   "Carrier_28_SpareSafetyInput(2_1)" AT %I1764.1 : Bool;   // SPARE SAFETY INPUT
   "Carrier_28_SpareSafetyInput(2_2)" AT %I1764.2 : Bool;   // SPARE SAFETY INPUT
   "Carrier_28_SpareSafetyInput(2_3)" AT %I1764.3 : Bool;   // SPARE SAFETY INPUT
   "Carrier_28_SpareSafetyInput(2_4)" AT %I1764.4 : Bool;   // SPARE SAFETY INPUT
   "Carrier_28_SpareSafetyInput(2_5)" AT %I1764.5 : Bool;   // SPARE SAFETY INPUT
   "Carrier_28_SpareSafetyInput(2_6)" AT %I1764.6 : Bool;   // SPARE SAFETY INPUT
   "Carrier_28_SpareSafetyInput(2_7)" AT %I1764.7 : Bool;   // SPARE SAFETY INPUT
   "Carrier_28_Slot3_SafetyOutput" AT %IW1675 : Word;   // SLOT 3 SAFETY OUTPUT WORD
   "Carrier_28_Crash_Detect_OK" AT %I1675.0 : Bool;   // CARRIER CRASH DETECT
   "Carrier_28_SpareSafetyOutput(3_1)" AT %I1675.1 : Bool;   // SPARE SAFETY OUTPUT
   "Carrier_28_SpareSafetyOutput(3_2)" AT %I1675.2 : Bool;   // SPARE SAFETY OUTPUT
   "Carrier_28_SpareSafetyOutput(3_3)" AT %I1675.3 : Bool;   // SPARE SAFETY OUTPUT
   "Carrier_28_SpareSafetyOutput(3_4)" AT %I1675.4 : Bool;   // SPARE SAFETY OUTPUT
   "Carrier_28_SpareSafetyOutput(3_5)" AT %I1675.5 : Bool;   // SPARE SAFETY OUTPUT
   "Carrier_28_SpareSafetyOutput(3_6)" AT %I1675.6 : Bool;   // SPARE SAFETY OUTPUT
   "Carrier_28_SpareSafetyOutput(3_7)" AT %I1675.7 : Bool;   // SPARE SAFETY OUTPUT
   "Carrier_28_Slot4_Input" AT %IW1766 : Word;   // SLOT 4 INPUT WORD
   "Carrier_28_480VPowerOn_MDCB1" AT %I1766.0 : Bool;   // 480 VAC POWER ON MDCB 1
   "Carrier_28_SpareInput(4_1)" AT %I1766.1 : Bool;   // SPARE INPUT
   "Carrier_28_SpareInput(4_2)" AT %I1766.2 : Bool;   // SPARE INPUT
   "Carrier_28_SitopSelectStatus" AT %I1766.3 : Bool;   // SITOP SELECT STATUS
   "Carrier_28_DCsupplyOnPSCB2" AT %I1766.4 : Bool;   // DC SUPPLY ON PSCB 2
   "Carrier_28_SpareInput(4_5)" AT %I1766.5 : Bool;   // SPARE INPUT
   "Carrier_28_SpareInput(4_6)" AT %I1766.6 : Bool;   // SPARE INPUT
   "Carrier_28_SpareInput(4_7)" AT %I1766.7 : Bool;   // SPARE INPUT
   "Carrier_28_PB1_ProdHoldLH" AT %I1767.0 : Bool;   // PB 1 PRODUCTION HOLD LH
   "Carrier_28_PB2_ResetLH" AT %I1767.1 : Bool;   // PB 2 RESET LH
   "Carrier_28_PB3_ProdHoldRH" AT %I1767.2 : Bool;   // PB 3 PRODUCTION HOLD RH
   "Carrier_28_PB4_ResetRH" AT %I1767.3 : Bool;   // PB 4 RESET RH
   "Carrier_28_SpareInput(4_14)" AT %I1767.4 : Bool;   // SPARE INPUT
   "Carrier_28_SpareInput(4_15)" AT %I1767.5 : Bool;   // SPARE INPUT
   "Carrier_28_SpareInput(4_16)" AT %I1767.6 : Bool;   // SPARE INPUT
   "Carrier_28_SpareInput(4_17)" AT %I1767.7 : Bool;   // SPARE INPUT
   "Carrier_28_Slot5_Output" AT %IW1768 : Word;   // SLOT 5 OUTPUT WORD
   "Carrier_28_IRD400_HMI_24VDC_ENABLE" AT %I1768.0 : Bool;   // IRD 400 PANEL HMI 24V DC POWER
   "Carrier_28_FaultLight_LH" AT %I1768.1 : Bool;   // FAULT LIGHT LH
   "Carrier_28_RunLight_LH" AT %I1768.2 : Bool;   // RUN LIGHT LH
   "Carrier_28_FaultLight_RH" AT %I1768.3 : Bool;   // FAULT LIGHT RH
   "Carrier_28_RunLight_RH" AT %I1768.4 : Bool;   // RUN LIGHT RH
   "Carrier_28_SpareOutput(5_5)" AT %I1768.5 : Bool;   // SPARE OUTPUT
   "Carrier_28_SpareOutput(5_6)" AT %I1768.6 : Bool;   // SPARE OUTPUT
   "Carrier_28_SpareOutput(5_7)" AT %I1768.7 : Bool;   // SPARE OUTPUT
   "Carrier_28_ActualSpeed" AT %IW1770 : Word;   // ACTUAL SPEED
   "Carrier_28_CarrierDriveAlarm" AT %IW1772 : Word;   // CARRIER DRIVE ALARM
   "Carrier_28_CarrierDriveWarning" AT %IW1774 : Word;   // CARRIER DRIVE WARNING
   "Carrier_29_Status" AT %IW1800 : Word;   // CARRIER STATUS WORD
   "Carrier_29_Status.0" AT %I1800.0 : Bool;   // HEARTBEAT
   "Carrier_29_Status.1" AT %I1800.1 : Bool;   // MANUAL
   "Carrier_29_Status.2" AT %I1800.2 : Bool;   // IN_AUTO
   "Carrier_29_Status.3" AT %I1800.3 : Bool;   // POSITIONING_COMPLETE
   "Carrier_29_Status.4" AT %I1800.4 : Bool;   // PRODUCTION HOLD
   "Carrier_29_Status.5" AT %I1800.5 : Bool;   // CARRIER MOVING FORWARD
   "Carrier_29_Status.6" AT %I1800.6 : Bool;   // CARRIER MOVING REVERSE
   "Carrier_29_Status.7" AT %I1800.7 : Bool;   // CARRIER FAULT
   "Carrier_29_Status.8" AT %I1801.0 : Bool;   // CRASH DETECT TRIPPED
   "Carrier_29_Status.9" AT %I1801.1 : Bool;
   "Carrier_29_Status.10" AT %I1801.2 : Bool;
   "Carrier_29_Status.11" AT %I1801.3 : Bool;
   "Carrier_29_Status.12" AT %I1801.4 : Bool;
   "Carrier_29_Status.13" AT %I1801.5 : Bool;
   "Carrier_29_Status.14" AT %I1801.6 : Bool;
   "Carrier_29_Status.15" AT %I1801.7 : Bool;
   "Carrier_29_SDCFaultCode" AT %IW1802 : Word;   // SDC FAULT CODE
   "Carrier_29_CarrierPosition" AT %ID1804 : DWord;   // CARRIER POSITION
   "Carrier_29_CarrierNumber" AT %IW1808 : Word;   // CARRIER NUMBER
   "Carrier_29_G120DControlWord" AT %IW1810 : Word;   // G120D_STW1_CONTROL
   "Carrier_29_G120DControlWord.0" AT %I1810.0 : Bool;   // Bit_00_ON
   "Carrier_29_G120DControlWord.1" AT %I1810.1 : Bool;   // Bit_01_AUS2_INH
   "Carrier_29_G120DControlWord.2" AT %I1810.2 : Bool;   // Bit_02_AUS3_STOP
   "Carrier_29_G120DControlWord.3" AT %I1810.3 : Bool;   // Bit_03_EN
   "Carrier_29_G120DControlWord.4" AT %I1810.4 : Bool;   // Bit_04_EN_RAMP
   "Carrier_29_G120DControlWord.5" AT %I1810.5 : Bool;   // Bit_05_START_RAMP
   "Carrier_29_G120DControlWord.6" AT %I1810.6 : Bool;   // Bit_06_SETPOINT
   "Carrier_29_G120DControlWord.7" AT %I1810.7 : Bool;   // Bit_07_RESET
   "Carrier_29_G120DControlWord.8" AT %I1811.0 : Bool;   // Bit_08_JOG_R
   "Carrier_29_G120DControlWord.9" AT %I1811.1 : Bool;   // Bit_09_JOG_L
   "Carrier_29_G120DControlWord.10" AT %I1811.2 : Bool;   // Bit_10_CONTR_PLC
   "Carrier_29_G120DControlWord.11" AT %I1811.3 : Bool;   // Bit_11_REVERSE
   "Carrier_29_G120DControlWord.12" AT %I1811.4 : Bool;   // Bit_12_BRAKE_RELEASE
   "Carrier_29_G120DControlWord.13" AT %I1811.5 : Bool;   // Bit_13_DDS
   "Carrier_29_G120DControlWord.14" AT %I1811.6 : Bool;   // Bit_14_DO0
   "Carrier_29_G120DControlWord.15" AT %I1811.7 : Bool;   // Bit_15_DO1
   "Carrier_29_G120DStatusWord" AT %IW1812 : Word;   // G120D_ZSW1_STATUS
   "Carrier_29_G120DStatusWord.0" AT %I1812.0 : Bool;   // Bit_00_READY_RUN
   "Carrier_29_G120DStatusWord.1" AT %I1812.1 : Bool;   // Bit_01_READY_ON
   "Carrier_29_G120DStatusWord.2" AT %I1812.2 : Bool;   // Bit_02_ENABLE
   "Carrier_29_G120DStatusWord.3" AT %I1812.3 : Bool;   // Bit_03_FAULT
   "Carrier_29_G120DStatusWord.4" AT %I1812.4 : Bool;   // Bit_04_OFF2
   "Carrier_29_G120DStatusWord.5" AT %I1812.5 : Bool;   // Bit_05_OFF3
   "Carrier_29_G120DStatusWord.6" AT %I1812.6 : Bool;   // Bit_06_LOCK_OUT
   "Carrier_29_G120DStatusWord.7" AT %I1812.7 : Bool;   // Bit_07_WARN
   "Carrier_29_G120DStatusWord.8" AT %I1813.0 : Bool;   // Bit_08_NO_DEVIATION
   "Carrier_29_G120DStatusWord.9" AT %I1813.1 : Bool;   // Bit_09_CONTR_PLC
   "Carrier_29_G120DStatusWord.10" AT %I1813.2 : Bool;   // Bit_10_F_MAX
   "Carrier_29_G120DStatusWord.11" AT %I1813.3 : Bool;   // Bit_11_LIMIT_REACHED
   "Carrier_29_G120DStatusWord.12" AT %I1813.4 : Bool;   // Bit_12_BRAKE_OPEN
   "Carrier_29_G120DStatusWord.13" AT %I1813.5 : Bool;   // Bit_13_NO_OVERTEMP
   "Carrier_29_G120DStatusWord.14" AT %I1813.6 : Bool;   // Bit_14_CW_CCW
   "Carrier_29_G120DStatusWord.15" AT %I1813.7 : Bool;   // Bit_15_OVERL
   "Carrier_29_Slot2_Input" AT %IW1814 : Word;   // SLOT 2 INPUT WORD
   "Carrier_29_CrashDetectSW" AT %I1814.0 : Bool;   // CRASH DETECT SW
   "Carrier_29_SpareSafetyInput(2_1)" AT %I1814.1 : Bool;   // SPARE SAFETY INPUT
   "Carrier_29_SpareSafetyInput(2_2)" AT %I1814.2 : Bool;   // SPARE SAFETY INPUT
   "Carrier_29_SpareSafetyInput(2_3)" AT %I1814.3 : Bool;   // SPARE SAFETY INPUT
   "Carrier_29_SpareSafetyInput(2_4)" AT %I1814.4 : Bool;   // SPARE SAFETY INPUT
   "Carrier_29_SpareSafetyInput(2_5)" AT %I1814.5 : Bool;   // SPARE SAFETY INPUT
   "Carrier_29_SpareSafetyInput(2_6)" AT %I1814.6 : Bool;   // SPARE SAFETY INPUT
   "Carrier_29_SpareSafetyInput(2_7)" AT %I1814.7 : Bool;   // SPARE SAFETY INPUT
   "Carrier_29_Slot3_SafetyOutput" AT %IW1815 : Word;   // SLOT 3 SAFETY OUTPUT WORD
   "Carrier_29_Crash_Detect_OK" AT %I1815.0 : Bool;   // CARRIER CRASH DETECT
   "Carrier_29_SpareSafetyOutput(3_1)" AT %I1815.1 : Bool;   // SPARE SAFETY OUTPUT
   "Carrier_29_SpareSafetyOutput(3_2)" AT %I1815.2 : Bool;   // SPARE SAFETY OUTPUT
   "Carrier_29_SpareSafetyOutput(3_3)" AT %I1815.3 : Bool;   // SPARE SAFETY OUTPUT
   "Carrier_29_SpareSafetyOutput(3_4)" AT %I1815.4 : Bool;   // SPARE SAFETY OUTPUT
   "Carrier_29_SpareSafetyOutput(3_5)" AT %I1815.5 : Bool;   // SPARE SAFETY OUTPUT
   "Carrier_29_SpareSafetyOutput(3_6)" AT %I1815.6 : Bool;   // SPARE SAFETY OUTPUT
   "Carrier_29_SpareSafetyOutput(3_7)" AT %I1815.7 : Bool;   // SPARE SAFETY OUTPUT
   "Carrier_29_Slot4_Input" AT %IW1816 : Word;   // SLOT 4 INPUT WORD
   "Carrier_29_480VPowerOn_MDCB1" AT %I1816.0 : Bool;   // 480 VAC POWER ON MDCB 1
   "Carrier_29_SpareInput(4_1)" AT %I1816.1 : Bool;   // SPARE INPUT
   "Carrier_29_SpareInput(4_2)" AT %I1816.2 : Bool;   // SPARE INPUT
   "Carrier_29_SitopSelectStatus" AT %I1816.3 : Bool;   // SITOP SELECT STATUS
   "Carrier_29_DCsupplyOnPSCB2" AT %I1816.4 : Bool;   // DC SUPPLY ON PSCB 2
   "Carrier_29_SpareInput(4_5)" AT %I1816.5 : Bool;   // SPARE INPUT
   "Carrier_29_SpareInput(4_6)" AT %I1816.6 : Bool;   // SPARE INPUT
   "Carrier_29_SpareInput(4_7)" AT %I1816.7 : Bool;   // SPARE INPUT
   "Carrier_29_PB1_ProdHoldLH" AT %I1817.0 : Bool;   // PB 1 PRODUCTION HOLD LH
   "Carrier_29_PB2_ResetLH" AT %I1817.1 : Bool;   // PB 2 RESET LH
   "Carrier_29_PB3_ProdHoldRH" AT %I1817.2 : Bool;   // PB 3 PRODUCTION HOLD RH
   "Carrier_29_PB4_ResetRH" AT %I1817.3 : Bool;   // PB 4 RESET RH
   "Carrier_29_SpareInput(4_14)" AT %I1817.4 : Bool;   // SPARE INPUT
   "Carrier_29_SpareInput(4_15)" AT %I1817.5 : Bool;   // SPARE INPUT
   "Carrier_29_SpareInput(4_16)" AT %I1817.6 : Bool;   // SPARE INPUT
   "Carrier_29_SpareInput(4_17)" AT %I1817.7 : Bool;   // SPARE INPUT
   "Carrier_29_Slot5_Output" AT %IW1818 : Word;   // SLOT 5 OUTPUT WORD
   "Carrier_29_IRD400_HMI_24VDC_ENABLE" AT %I1818.0 : Bool;   // IRD 400 PANEL HMI 24V DC POWER
   "Carrier_29_FaultLight_LH" AT %I1818.1 : Bool;   // FAULT LIGHT LH
   "Carrier_29_RunLight_LH" AT %I1818.2 : Bool;   // RUN LIGHT LH
   "Carrier_29_FaultLight_RH" AT %I1818.3 : Bool;   // FAULT LIGHT RH
   "Carrier_29_RunLight_RH" AT %I1818.4 : Bool;   // RUN LIGHT RH
   "Carrier_29_SpareOutput(5_5)" AT %I1818.5 : Bool;   // SPARE OUTPUT
   "Carrier_29_SpareOutput(5_6)" AT %I1818.6 : Bool;   // SPARE OUTPUT
   "Carrier_29_SpareOutput(5_7)" AT %I1818.7 : Bool;   // SPARE OUTPUT
   "Carrier_29_ActualSpeed" AT %IW1820 : Word;   // ACTUAL SPEED
   "Carrier_29_CarrierDriveAlarm" AT %IW1822 : Word;   // CARRIER DRIVE ALARM
   "Carrier_29_CarrierDriveWarning" AT %IW1824 : Word;   // CARRIER DRIVE WARNING
   "Carrier_30_Status" AT %IW1850 : Word;   // CARRIER STATUS WORD
   "Carrier_30_Status.0" AT %I1850.0 : Bool;   // HEARTBEAT
   "Carrier_30_Status.1" AT %I1850.1 : Bool;   // MANUAL
   "Carrier_30_Status.2" AT %I1850.2 : Bool;   // IN_AUTO
   "Carrier_30_Status.3" AT %I1850.3 : Bool;   // POSITIONING_COMPLETE
   "Carrier_30_Status.4" AT %I1850.4 : Bool;   // PRODUCTION HOLD
   "Carrier_30_Status.5" AT %I1850.5 : Bool;   // CARRIER MOVING FORWARD
   "Carrier_30_Status.6" AT %I1850.6 : Bool;   // CARRIER MOVING REVERSE
   "Carrier_30_Status.7" AT %I1850.7 : Bool;   // CARRIER FAULT
   "Carrier_30_Status.8" AT %I1851.0 : Bool;   // CRASH DETECT TRIPPED
   "Carrier_30_Status.9" AT %I1851.1 : Bool;
   "Carrier_30_Status.10" AT %I1851.2 : Bool;
   "Carrier_30_Status.11" AT %I1851.3 : Bool;
   "Carrier_30_Status.12" AT %I1851.4 : Bool;
   "Carrier_30_Status.13" AT %I1851.5 : Bool;
   "Carrier_30_Status.14" AT %I1851.6 : Bool;
   "Carrier_30_Status.15" AT %I1851.7 : Bool;
   "Carrier_30_SDCFaultCode" AT %IW1852 : Word;   // SDC FAULT CODE
   "Carrier_30_CarrierPosition" AT %ID1854 : DWord;   // CARRIER POSITION
   "Carrier_30_CarrierNumber" AT %IW1858 : Word;   // CARRIER NUMBER
   "Carrier_30_G120DControlWord" AT %IW1860 : Word;   // G120D_STW1_CONTROL
   "Carrier_30_G120DControlWord.0" AT %I1860.0 : Bool;   // Bit_00_ON
   "Carrier_30_G120DControlWord.1" AT %I1860.1 : Bool;   // Bit_01_AUS2_INH
   "Carrier_30_G120DControlWord.2" AT %I1860.2 : Bool;   // Bit_02_AUS3_STOP
   "Carrier_30_G120DControlWord.3" AT %I1860.3 : Bool;   // Bit_03_EN
   "Carrier_30_G120DControlWord.4" AT %I1860.4 : Bool;   // Bit_04_EN_RAMP
   "Carrier_30_G120DControlWord.5" AT %I1860.5 : Bool;   // Bit_05_START_RAMP
   "Carrier_30_G120DControlWord.6" AT %I1860.6 : Bool;   // Bit_06_SETPOINT
   "Carrier_30_G120DControlWord.7" AT %I1860.7 : Bool;   // Bit_07_RESET
   "Carrier_30_G120DControlWord.8" AT %I1861.0 : Bool;   // Bit_08_JOG_R
   "Carrier_30_G120DControlWord.9" AT %I1861.1 : Bool;   // Bit_09_JOG_L
   "Carrier_30_G120DControlWord.10" AT %I1861.2 : Bool;   // Bit_10_CONTR_PLC
   "Carrier_30_G120DControlWord.11" AT %I1861.3 : Bool;   // Bit_11_REVERSE
   "Carrier_30_G120DControlWord.12" AT %I1861.4 : Bool;   // Bit_12_BRAKE_RELEASE
   "Carrier_30_G120DControlWord.13" AT %I1861.5 : Bool;   // Bit_13_DDS
   "Carrier_30_G120DControlWord.14" AT %I1861.6 : Bool;   // Bit_14_DO0
   "Carrier_30_G120DControlWord.15" AT %I1861.7 : Bool;   // Bit_15_DO1
   "Carrier_30_G120DStatusWord" AT %IW1862 : Word;   // G120D_ZSW1_STATUS
   "Carrier_30_G120DStatusWord.0" AT %I1862.0 : Bool;   // Bit_00_READY_RUN
   "Carrier_30_G120DStatusWord.1" AT %I1862.1 : Bool;   // Bit_01_READY_ON
   "Carrier_30_G120DStatusWord.2" AT %I1862.2 : Bool;   // Bit_02_ENABLE
   "Carrier_30_G120DStatusWord.3" AT %I1862.3 : Bool;   // Bit_03_FAULT
   "Carrier_30_G120DStatusWord.4" AT %I1862.4 : Bool;   // Bit_04_OFF2
   "Carrier_30_G120DStatusWord.5" AT %I1862.5 : Bool;   // Bit_05_OFF3
   "Carrier_30_G120DStatusWord.6" AT %I1862.6 : Bool;   // Bit_06_LOCK_OUT
   "Carrier_30_G120DStatusWord.7" AT %I1862.7 : Bool;   // Bit_07_WARN
   "Carrier_30_G120DStatusWord.8" AT %I1863.0 : Bool;   // Bit_08_NO_DEVIATION
   "Carrier_30_G120DStatusWord.9" AT %I1863.1 : Bool;   // Bit_09_CONTR_PLC
   "Carrier_30_G120DStatusWord.10" AT %I1863.2 : Bool;   // Bit_10_F_MAX
   "Carrier_30_G120DStatusWord.11" AT %I1863.3 : Bool;   // Bit_11_LIMIT_REACHED
   "Carrier_30_G120DStatusWord.12" AT %I1863.4 : Bool;   // Bit_12_BRAKE_OPEN
   "Carrier_30_G120DStatusWord.13" AT %I1863.5 : Bool;   // Bit_13_NO_OVERTEMP
   "Carrier_30_G120DStatusWord.14" AT %I1863.6 : Bool;   // Bit_14_CW_CCW
   "Carrier_30_G120DStatusWord.15" AT %I1863.7 : Bool;   // Bit_15_OVERL
   "Carrier_30_Slot2_Input" AT %IW1864 : Word;   // SLOT 2 INPUT WORD
   "Carrier_30_CrashDetectSW" AT %I1864.0 : Bool;   // CRASH DETECT SW
   "Carrier_30_SpareSafetyInput(2_1)" AT %I1864.1 : Bool;   // SPARE SAFETY INPUT
   "Carrier_30_SpareSafetyInput(2_2)" AT %I1864.2 : Bool;   // SPARE SAFETY INPUT
   "Carrier_30_SpareSafetyInput(2_3)" AT %I1864.3 : Bool;   // SPARE SAFETY INPUT
   "Carrier_30_SpareSafetyInput(2_4)" AT %I1864.4 : Bool;   // SPARE SAFETY INPUT
   "Carrier_30_SpareSafetyInput(2_5)" AT %I1864.5 : Bool;   // SPARE SAFETY INPUT
   "Carrier_30_SpareSafetyInput(2_6)" AT %I1864.6 : Bool;   // SPARE SAFETY INPUT
   "Carrier_30_SpareSafetyInput(2_7)" AT %I1864.7 : Bool;   // SPARE SAFETY INPUT
   "Carrier_30_Slot3_SafetyOutput" AT %IW1685 : Word;   // SLOT 3 SAFETY OUTPUT WORD
   "Carrier_30_Crash_Detect_OK" AT %I1685.0 : Bool;   // CARRIER CRASH DETECT
   "Carrier_30_SpareSafetyOutput(3_1)" AT %I1685.1 : Bool;   // SPARE SAFETY OUTPUT
   "Carrier_30_SpareSafetyOutput(3_2)" AT %I1685.2 : Bool;   // SPARE SAFETY OUTPUT
   "Carrier_30_SpareSafetyOutput(3_3)" AT %I1685.3 : Bool;   // SPARE SAFETY OUTPUT
   "Carrier_30_SpareSafetyOutput(3_4)" AT %I1685.4 : Bool;   // SPARE SAFETY OUTPUT
   "Carrier_30_SpareSafetyOutput(3_5)" AT %I1685.5 : Bool;   // SPARE SAFETY OUTPUT
   "Carrier_30_SpareSafetyOutput(3_6)" AT %I1685.6 : Bool;   // SPARE SAFETY OUTPUT
   "Carrier_30_SpareSafetyOutput(3_7)" AT %I1685.7 : Bool;   // SPARE SAFETY OUTPUT
   "Carrier_30_Slot4_Input" AT %IW1866 : Word;   // SLOT 4 INPUT WORD
   "Carrier_30_480VPowerOn_MDCB1" AT %I1866.0 : Bool;   // 480 VAC POWER ON MDCB 1
   "Carrier_30_SpareInput(4_1)" AT %I1866.1 : Bool;   // SPARE INPUT
   "Carrier_30_SpareInput(4_2)" AT %I1866.2 : Bool;   // SPARE INPUT
   "Carrier_30_SitopSelectStatus" AT %I1866.3 : Bool;   // SITOP SELECT STATUS
   "Carrier_30_DCsupplyOnPSCB2" AT %I1866.4 : Bool;   // DC SUPPLY ON PSCB 2
   "Carrier_30_SpareInput(4_5)" AT %I1866.5 : Bool;   // SPARE INPUT
   "Carrier_30_SpareInput(4_6)" AT %I1866.6 : Bool;   // SPARE INPUT
   "Carrier_30_SpareInput(4_7)" AT %I1866.7 : Bool;   // SPARE INPUT
   "Carrier_30_PB1_ProdHoldLH" AT %I1867.0 : Bool;   // PB 1 PRODUCTION HOLD LH
   "Carrier_30_PB2_ResetLH" AT %I1867.1 : Bool;   // PB 2 RESET LH
   "Carrier_30_PB3_ProdHoldRH" AT %I1867.2 : Bool;   // PB 3 PRODUCTION HOLD RH
   "Carrier_30_PB4_ResetRH" AT %I1867.3 : Bool;   // PB 4 RESET RH
   "Carrier_30_SpareInput(4_14)" AT %I1867.4 : Bool;   // SPARE INPUT
   "Carrier_30_SpareInput(4_15)" AT %I1867.5 : Bool;   // SPARE INPUT
   "Carrier_30_SpareInput(4_16)" AT %I1867.6 : Bool;   // SPARE INPUT
   "Carrier_30_SpareInput(4_17)" AT %I1867.7 : Bool;   // SPARE INPUT
   "Carrier_30_Slot5_Output" AT %IW1868 : Word;   // SLOT 5 OUTPUT WORD
   "Carrier_30_IRD400_HMI_24VDC_ENABLE" AT %I1868.0 : Bool;   // IRD 400 PANEL HMI 24V DC POWER
   "Carrier_30_FaultLight_LH" AT %I1868.1 : Bool;   // FAULT LIGHT LH
   "Carrier_30_RunLight_LH" AT %I1868.2 : Bool;   // RUN LIGHT LH
   "Carrier_30_FaultLight_RH" AT %I1868.3 : Bool;   // FAULT LIGHT RH
   "Carrier_30_RunLight_RH" AT %I1868.4 : Bool;   // RUN LIGHT RH
   "Carrier_30_SpareOutput(5_5)" AT %I1868.5 : Bool;   // SPARE OUTPUT
   "Carrier_30_SpareOutput(5_6)" AT %I1868.6 : Bool;   // SPARE OUTPUT
   "Carrier_30_SpareOutput(5_7)" AT %I1868.7 : Bool;   // SPARE OUTPUT
   "Carrier_30_ActualSpeed" AT %IW1870 : Word;   // ACTUAL SPEED
   "Carrier_30_CarrierDriveAlarm" AT %IW1872 : Word;   // CARRIER DRIVE ALARM
   "Carrier_30_CarrierDriveWarning" AT %IW1874 : Word;   // CARRIER DRIVE WARNING
   "Carrier_31_Status" AT %IW1900 : Word;   // CARRIER STATUS WORD
   "Carrier_31_Status.0" AT %I1900.0 : Bool;   // HEARTBEAT
   "Carrier_31_Status.1" AT %I1900.1 : Bool;   // MANUAL
   "Carrier_31_Status.2" AT %I1900.2 : Bool;   // IN_AUTO
   "Carrier_31_Status.3" AT %I1900.3 : Bool;   // POSITIONING_COMPLETE
   "Carrier_31_Status.4" AT %I1900.4 : Bool;   // PRODUCTION HOLD
   "Carrier_31_Status.5" AT %I1900.5 : Bool;   // CARRIER MOVING FORWARD
   "Carrier_31_Status.6" AT %I1900.6 : Bool;   // CARRIER MOVING REVERSE
   "Carrier_31_Status.7" AT %I1900.7 : Bool;   // CARRIER FAULT
   "Carrier_31_Status.8" AT %I1901.0 : Bool;   // CRASH DETECT TRIPPED
   "Carrier_31_Status.9" AT %I1901.1 : Bool;
   "Carrier_31_Status.10" AT %I1901.2 : Bool;
   "Carrier_31_Status.11" AT %I1901.3 : Bool;
   "Carrier_31_Status.12" AT %I1901.4 : Bool;
   "Carrier_31_Status.13" AT %I1901.5 : Bool;
   "Carrier_31_Status.14" AT %I1901.6 : Bool;
   "Carrier_31_Status.15" AT %I1901.7 : Bool;
   "Carrier_31_SDCFaultCode" AT %IW1902 : Word;   // SDC FAULT CODE
   "Carrier_31_CarrierPosition" AT %ID1904 : DWord;   // CARRIER POSITION
   "Carrier_31_CarrierNumber" AT %IW1908 : Word;   // CARRIER NUMBER
   "Carrier_31_G120DControlWord" AT %IW1910 : Word;   // G120D_STW1_CONTROL
   "Carrier_31_G120DControlWord.0" AT %I1910.0 : Bool;   // Bit_00_ON
   "Carrier_31_G120DControlWord.1" AT %I1910.1 : Bool;   // Bit_01_AUS2_INH
   "Carrier_31_G120DControlWord.2" AT %I1910.2 : Bool;   // Bit_02_AUS3_STOP
   "Carrier_31_G120DControlWord.3" AT %I1910.3 : Bool;   // Bit_03_EN
   "Carrier_31_G120DControlWord.4" AT %I1910.4 : Bool;   // Bit_04_EN_RAMP
   "Carrier_31_G120DControlWord.5" AT %I1910.5 : Bool;   // Bit_05_START_RAMP
   "Carrier_31_G120DControlWord.6" AT %I1910.6 : Bool;   // Bit_06_SETPOINT
   "Carrier_31_G120DControlWord.7" AT %I1910.7 : Bool;   // Bit_07_RESET
   "Carrier_31_G120DControlWord.8" AT %I1911.0 : Bool;   // Bit_08_JOG_R
   "Carrier_31_G120DControlWord.9" AT %I1911.1 : Bool;   // Bit_09_JOG_L
   "Carrier_31_G120DControlWord.10" AT %I1911.2 : Bool;   // Bit_10_CONTR_PLC
   "Carrier_31_G120DControlWord.11" AT %I1911.3 : Bool;   // Bit_11_REVERSE
   "Carrier_31_G120DControlWord.12" AT %I1911.4 : Bool;   // Bit_12_BRAKE_RELEASE
   "Carrier_31_G120DControlWord.13" AT %I1911.5 : Bool;   // Bit_13_DDS
   "Carrier_31_G120DControlWord.14" AT %I1911.6 : Bool;   // Bit_14_DO0
   "Carrier_31_G120DControlWord.15" AT %I1911.7 : Bool;   // Bit_15_DO1
   "Carrier_31_G120DStatusWord" AT %IW1912 : Word;   // G120D_ZSW1_STATUS
   "Carrier_31_G120DStatusWord.0" AT %I1912.0 : Bool;   // Bit_00_READY_RUN
   "Carrier_31_G120DStatusWord.1" AT %I1912.1 : Bool;   // Bit_01_READY_ON
   "Carrier_31_G120DStatusWord.2" AT %I1912.2 : Bool;   // Bit_02_ENABLE
   "Carrier_31_G120DStatusWord.3" AT %I1912.3 : Bool;   // Bit_03_FAULT
   "Carrier_31_G120DStatusWord.4" AT %I1912.4 : Bool;   // Bit_04_OFF2
   "Carrier_31_G120DStatusWord.5" AT %I1912.5 : Bool;   // Bit_05_OFF3
   "Carrier_31_G120DStatusWord.6" AT %I1912.6 : Bool;   // Bit_06_LOCK_OUT
   "Carrier_31_G120DStatusWord.7" AT %I1912.7 : Bool;   // Bit_07_WARN
   "Carrier_31_G120DStatusWord.8" AT %I1913.0 : Bool;   // Bit_08_NO_DEVIATION
   "Carrier_31_G120DStatusWord.9" AT %I1913.1 : Bool;   // Bit_09_CONTR_PLC
   "Carrier_31_G120DStatusWord.10" AT %I1913.2 : Bool;   // Bit_10_F_MAX
   "Carrier_31_G120DStatusWord.11" AT %I1913.3 : Bool;   // Bit_11_LIMIT_REACHED
   "Carrier_31_G120DStatusWord.12" AT %I1913.4 : Bool;   // Bit_12_BRAKE_OPEN
   "Carrier_31_G120DStatusWord.13" AT %I1913.5 : Bool;   // Bit_13_NO_OVERTEMP
   "Carrier_31_G120DStatusWord.14" AT %I1913.6 : Bool;   // Bit_14_CW_CCW
   "Carrier_31_G120DStatusWord.15" AT %I1913.7 : Bool;   // Bit_15_OVERL
   "Carrier_31_Slot2_Input" AT %IW1914 : Word;   // SLOT 2 INPUT WORD
   "Carrier_31_CrashDetectSW" AT %I1914.0 : Bool;   // CRASH DETECT SW
   "Carrier_31_SpareSafetyInput(2_1)" AT %I1914.1 : Bool;   // SPARE SAFETY INPUT
   "Carrier_31_SpareSafetyInput(2_2)" AT %I1914.2 : Bool;   // SPARE SAFETY INPUT
   "Carrier_31_SpareSafetyInput(2_3)" AT %I1914.3 : Bool;   // SPARE SAFETY INPUT
   "Carrier_31_SpareSafetyInput(2_4)" AT %I1914.4 : Bool;   // SPARE SAFETY INPUT
   "Carrier_31_SpareSafetyInput(2_5)" AT %I1914.5 : Bool;   // SPARE SAFETY INPUT
   "Carrier_31_SpareSafetyInput(2_6)" AT %I1914.6 : Bool;   // SPARE SAFETY INPUT
   "Carrier_31_SpareSafetyInput(2_7)" AT %I1914.7 : Bool;   // SPARE SAFETY INPUT
   "Carrier_31_Slot3_SafetyOutput" AT %IW1915 : Word;   // SLOT 3 SAFETY OUTPUT WORD
   "Carrier_31_Crash_Detect_OK" AT %I1915.0 : Bool;   // CARRIER CRASH DETECT
   "Carrier_31_SpareSafetyOutput(3_1)" AT %I1915.1 : Bool;   // SPARE SAFETY OUTPUT
   "Carrier_31_SpareSafetyOutput(3_2)" AT %I1915.2 : Bool;   // SPARE SAFETY OUTPUT
   "Carrier_31_SpareSafetyOutput(3_3)" AT %I1915.3 : Bool;   // SPARE SAFETY OUTPUT
   "Carrier_31_SpareSafetyOutput(3_4)" AT %I1915.4 : Bool;   // SPARE SAFETY OUTPUT
   "Carrier_31_SpareSafetyOutput(3_5)" AT %I1915.5 : Bool;   // SPARE SAFETY OUTPUT
   "Carrier_31_SpareSafetyOutput(3_6)" AT %I1915.6 : Bool;   // SPARE SAFETY OUTPUT
   "Carrier_31_SpareSafetyOutput(3_7)" AT %I1915.7 : Bool;   // SPARE SAFETY OUTPUT
   "Carrier_31_Slot4_Input" AT %IW1916 : Word;   // SLOT 4 INPUT WORD
   "Carrier_31_480VPowerOn_MDCB1" AT %I1916.0 : Bool;   // 480 VAC POWER ON MDCB 1
   "Carrier_31_SpareInput(4_1)" AT %I1916.1 : Bool;   // SPARE INPUT
   "Carrier_31_SpareInput(4_2)" AT %I1916.2 : Bool;   // SPARE INPUT
   "Carrier_31_SitopSelectStatus" AT %I1916.3 : Bool;   // SITOP SELECT STATUS
   "Carrier_31_DCsupplyOnPSCB2" AT %I1916.4 : Bool;   // DC SUPPLY ON PSCB 2
   "Carrier_31_SpareInput(4_5)" AT %I1916.5 : Bool;   // SPARE INPUT
   "Carrier_31_SpareInput(4_6)" AT %I1916.6 : Bool;   // SPARE INPUT
   "Carrier_31_SpareInput(4_7)" AT %I1916.7 : Bool;   // SPARE INPUT
   "Carrier_31_PB1_ProdHoldLH" AT %I1917.0 : Bool;   // PB 1 PRODUCTION HOLD LH
   "Carrier_31_PB2_ResetLH" AT %I1917.1 : Bool;   // PB 2 RESET LH
   "Carrier_31_PB3_ProdHoldRH" AT %I1917.2 : Bool;   // PB 3 PRODUCTION HOLD RH
   "Carrier_31_PB4_ResetRH" AT %I1917.3 : Bool;   // PB 4 RESET RH
   "Carrier_31_SpareInput(4_14)" AT %I1917.4 : Bool;   // SPARE INPUT
   "Carrier_31_SpareInput(4_15)" AT %I1917.5 : Bool;   // SPARE INPUT
   "Carrier_31_SpareInput(4_16)" AT %I1917.6 : Bool;   // SPARE INPUT
   "Carrier_31_SpareInput(4_17)" AT %I1917.7 : Bool;   // SPARE INPUT
   "Carrier_31_Slot5_Output" AT %IW1918 : Word;   // SLOT 5 OUTPUT WORD
   "Carrier_31_IRD400_HMI_24VDC_ENABLE" AT %I1918.0 : Bool;   // IRD 400 PANEL HMI 24V DC POWER
   "Carrier_31_FaultLight_LH" AT %I1918.1 : Bool;   // FAULT LIGHT LH
   "Carrier_31_RunLight_LH" AT %I1918.2 : Bool;   // RUN LIGHT LH
   "Carrier_31_FaultLight_RH" AT %I1918.3 : Bool;   // FAULT LIGHT RH
   "Carrier_31_RunLight_RH" AT %I1918.4 : Bool;   // RUN LIGHT RH
   "Carrier_31_SpareOutput(5_5)" AT %I1918.5 : Bool;   // SPARE OUTPUT
   "Carrier_31_SpareOutput(5_6)" AT %I1918.6 : Bool;   // SPARE OUTPUT
   "Carrier_31_SpareOutput(5_7)" AT %I1918.7 : Bool;   // SPARE OUTPUT
   "Carrier_31_ActualSpeed" AT %IW1920 : Word;   // ACTUAL SPEED
   "Carrier_31_CarrierDriveAlarm" AT %IW1922 : Word;   // CARRIER DRIVE ALARM
   "Carrier_31_CarrierDriveWarning" AT %IW1924 : Word;   // CARRIER DRIVE WARNING
   "Carrier_32_Status" AT %IW1950 : Word;   // CARRIER STATUS WORD
   "Carrier_32_Status.0" AT %I1950.0 : Bool;   // HEARTBEAT
   "Carrier_32_Status.1" AT %I1950.1 : Bool;   // MANUAL
   "Carrier_32_Status.2" AT %I1950.2 : Bool;   // IN_AUTO
   "Carrier_32_Status.3" AT %I1950.3 : Bool;   // POSITIONING_COMPLETE
   "Carrier_32_Status.4" AT %I1950.4 : Bool;   // PRODUCTION HOLD
   "Carrier_32_Status.5" AT %I1950.5 : Bool;   // CARRIER MOVING FORWARD
   "Carrier_32_Status.6" AT %I1950.6 : Bool;   // CARRIER MOVING REVERSE
   "Carrier_32_Status.7" AT %I1950.7 : Bool;   // CARRIER FAULT
   "Carrier_32_Status.8" AT %I1951.0 : Bool;   // CRASH DETECT TRIPPED
   "Carrier_32_Status.9" AT %I1951.1 : Bool;
   "Carrier_32_Status.10" AT %I1951.2 : Bool;
   "Carrier_32_Status.11" AT %I1951.3 : Bool;
   "Carrier_32_Status.12" AT %I1951.4 : Bool;
   "Carrier_32_Status.13" AT %I1951.5 : Bool;
   "Carrier_32_Status.14" AT %I1951.6 : Bool;
   "Carrier_32_Status.15" AT %I1951.7 : Bool;
   "Carrier_32_SDCFaultCode" AT %IW1952 : Word;   // SDC FAULT CODE
   "Carrier_32_CarrierPosition" AT %ID1954 : DWord;   // CARRIER POSITION
   "Carrier_32_CarrierNumber" AT %IW1958 : Word;   // CARRIER NUMBER
   "Carrier_32_G120DControlWord" AT %IW1960 : Word;   // G120D_STW1_CONTROL
   "Carrier_32_G120DControlWord.0" AT %I1960.0 : Bool;   // Bit_00_ON
   "Carrier_32_G120DControlWord.1" AT %I1960.1 : Bool;   // Bit_01_AUS2_INH
   "Carrier_32_G120DControlWord.2" AT %I1960.2 : Bool;   // Bit_02_AUS3_STOP
   "Carrier_32_G120DControlWord.3" AT %I1960.3 : Bool;   // Bit_03_EN
   "Carrier_32_G120DControlWord.4" AT %I1960.4 : Bool;   // Bit_04_EN_RAMP
   "Carrier_32_G120DControlWord.5" AT %I1960.5 : Bool;   // Bit_05_START_RAMP
   "Carrier_32_G120DControlWord.6" AT %I1960.6 : Bool;   // Bit_06_SETPOINT
   "Carrier_32_G120DControlWord.7" AT %I1960.7 : Bool;   // Bit_07_RESET
   "Carrier_32_G120DControlWord.8" AT %I1961.0 : Bool;   // Bit_08_JOG_R
   "Carrier_32_G120DControlWord.9" AT %I1961.1 : Bool;   // Bit_09_JOG_L
   "Carrier_32_G120DControlWord.10" AT %I1961.2 : Bool;   // Bit_10_CONTR_PLC
   "Carrier_32_G120DControlWord.11" AT %I1961.3 : Bool;   // Bit_11_REVERSE
   "Carrier_32_G120DControlWord.12" AT %I1961.4 : Bool;   // Bit_12_BRAKE_RELEASE
   "Carrier_32_G120DControlWord.13" AT %I1961.5 : Bool;   // Bit_13_DDS
   "Carrier_32_G120DControlWord.14" AT %I1961.6 : Bool;   // Bit_14_DO0
   "Carrier_32_G120DControlWord.15" AT %I1961.7 : Bool;   // Bit_15_DO1
   "Carrier_32_G120DStatusWord" AT %IW1962 : Word;   // G120D_ZSW1_STATUS
   "Carrier_32_G120DStatusWord.0" AT %I1962.0 : Bool;   // Bit_00_READY_RUN
   "Carrier_32_G120DStatusWord.1" AT %I1962.1 : Bool;   // Bit_01_READY_ON
   "Carrier_32_G120DStatusWord.2" AT %I1962.2 : Bool;   // Bit_02_ENABLE
   "Carrier_32_G120DStatusWord.3" AT %I1962.3 : Bool;   // Bit_03_FAULT
   "Carrier_32_G120DStatusWord.4" AT %I1962.4 : Bool;   // Bit_04_OFF2
   "Carrier_32_G120DStatusWord.5" AT %I1962.5 : Bool;   // Bit_05_OFF3
   "Carrier_32_G120DStatusWord.6" AT %I1962.6 : Bool;   // Bit_06_LOCK_OUT
   "Carrier_32_G120DStatusWord.7" AT %I1962.7 : Bool;   // Bit_07_WARN
   "Carrier_32_G120DStatusWord.8" AT %I1963.0 : Bool;   // Bit_08_NO_DEVIATION
   "Carrier_32_G120DStatusWord.9" AT %I1963.1 : Bool;   // Bit_09_CONTR_PLC
   "Carrier_32_G120DStatusWord.10" AT %I1963.2 : Bool;   // Bit_10_F_MAX
   "Carrier_32_G120DStatusWord.11" AT %I1963.3 : Bool;   // Bit_11_LIMIT_REACHED
   "Carrier_32_G120DStatusWord.12" AT %I1963.4 : Bool;   // Bit_12_BRAKE_OPEN
   "Carrier_32_G120DStatusWord.13" AT %I1963.5 : Bool;   // Bit_13_NO_OVERTEMP
   "Carrier_32_G120DStatusWord.14" AT %I1963.6 : Bool;   // Bit_14_CW_CCW
   "Carrier_32_G120DStatusWord.15" AT %I1963.7 : Bool;   // Bit_15_OVERL
   "Carrier_32_Slot2_Input" AT %IW1964 : Word;   // SLOT 2 INPUT WORD
   "Carrier_32_CrashDetectSW" AT %I1964.0 : Bool;   // CRASH DETECT SW
   "Carrier_32_SpareSafetyInput(2_1)" AT %I1964.1 : Bool;   // SPARE SAFETY INPUT
   "Carrier_32_SpareSafetyInput(2_2)" AT %I1964.2 : Bool;   // SPARE SAFETY INPUT
   "Carrier_32_SpareSafetyInput(2_3)" AT %I1964.3 : Bool;   // SPARE SAFETY INPUT
   "Carrier_32_SpareSafetyInput(2_4)" AT %I1964.4 : Bool;   // SPARE SAFETY INPUT
   "Carrier_32_SpareSafetyInput(2_5)" AT %I1964.5 : Bool;   // SPARE SAFETY INPUT
   "Carrier_32_SpareSafetyInput(2_6)" AT %I1964.6 : Bool;   // SPARE SAFETY INPUT
   "Carrier_32_SpareSafetyInput(2_7)" AT %I1964.7 : Bool;   // SPARE SAFETY INPUT
   "Carrier_32_Slot3_SafetyOutput" AT %IW1965 : Word;   // SLOT 3 SAFETY OUTPUT WORD
   "Carrier_32_Crash_Detect_OK" AT %I1965.0 : Bool;   // CARRIER CRASH DETECT
   "Carrier_32_SpareSafetyOutput(3_1)" AT %I1965.1 : Bool;   // SPARE SAFETY OUTPUT
   "Carrier_32_SpareSafetyOutput(3_2)" AT %I1965.2 : Bool;   // SPARE SAFETY OUTPUT
   "Carrier_32_SpareSafetyOutput(3_3)" AT %I1965.3 : Bool;   // SPARE SAFETY OUTPUT
   "Carrier_32_SpareSafetyOutput(3_4)" AT %I1965.4 : Bool;   // SPARE SAFETY OUTPUT
   "Carrier_32_SpareSafetyOutput(3_5)" AT %I1965.5 : Bool;   // SPARE SAFETY OUTPUT
   "Carrier_32_SpareSafetyOutput(3_6)" AT %I1965.6 : Bool;   // SPARE SAFETY OUTPUT
   "Carrier_32_SpareSafetyOutput(3_7)" AT %I1965.7 : Bool;   // SPARE SAFETY OUTPUT
   "Carrier_32_Slot4_Input" AT %IW1966 : Word;   // SLOT 4 INPUT WORD
   "Carrier_32_480VPowerOn_MDCB1" AT %I1966.0 : Bool;   // 480 VAC POWER ON MDCB 1
   "Carrier_32_SpareInput(4_1)" AT %I1966.1 : Bool;   // SPARE INPUT
   "Carrier_32_SpareInput(4_2)" AT %I1966.2 : Bool;   // SPARE INPUT
   "Carrier_32_SitopSelectStatus" AT %I1966.3 : Bool;   // SITOP SELECT STATUS
   "Carrier_32_DCsupplyOnPSCB2" AT %I1966.4 : Bool;   // DC SUPPLY ON PSCB 2
   "Carrier_32_SpareInput(4_5)" AT %I1966.5 : Bool;   // SPARE INPUT
   "Carrier_32_SpareInput(4_6)" AT %I1966.6 : Bool;   // SPARE INPUT
   "Carrier_32_SpareInput(4_7)" AT %I1966.7 : Bool;   // SPARE INPUT
   "Carrier_32_PB1_ProdHoldLH" AT %I1967.0 : Bool;   // PB 1 PRODUCTION HOLD LH
   "Carrier_32_PB2_ResetLH" AT %I1967.1 : Bool;   // PB 2 RESET LH
   "Carrier_32_PB3_ProdHoldRH" AT %I1967.2 : Bool;   // PB 3 PRODUCTION HOLD RH
   "Carrier_32_PB4_ResetRH" AT %I1967.3 : Bool;   // PB 4 RESET RH
   "Carrier_32_SpareInput(4_14)" AT %I1967.4 : Bool;   // SPARE INPUT
   "Carrier_32_SpareInput(4_15)" AT %I1967.5 : Bool;   // SPARE INPUT
   "Carrier_32_SpareInput(4_16)" AT %I1967.6 : Bool;   // SPARE INPUT
   "Carrier_32_SpareInput(4_17)" AT %I1967.7 : Bool;   // SPARE INPUT
   "Carrier_32_Slot5_Output" AT %IW1968 : Word;   // SLOT 5 OUTPUT WORD
   "Carrier_32_IRD400_HMI_24VDC_ENABLE" AT %I1968.0 : Bool;   // IRD 400 PANEL HMI 24V DC POWER
   "Carrier_32_FaultLight_LH" AT %I1968.1 : Bool;   // FAULT LIGHT LH
   "Carrier_32_RunLight_LH" AT %I1968.2 : Bool;   // RUN LIGHT LH
   "Carrier_32_FaultLight_RH" AT %I1968.3 : Bool;   // FAULT LIGHT RH
   "Carrier_32_RunLight_RH" AT %I1968.4 : Bool;   // RUN LIGHT RH
   "Carrier_32_SpareOutput(5_5)" AT %I1968.5 : Bool;   // SPARE OUTPUT
   "Carrier_32_SpareOutput(5_6)" AT %I1968.6 : Bool;   // SPARE OUTPUT
   "Carrier_32_SpareOutput(5_7)" AT %I1968.7 : Bool;   // SPARE OUTPUT
   "Carrier_32_ActualSpeed" AT %IW1970 : Word;   // ACTUAL SPEED
   "Carrier_32_CarrierDriveAlarm" AT %IW1972 : Word;   // CARRIER DRIVE ALARM
   "Carrier_32_CarrierDriveWarning" AT %IW1974 : Word;   // CARRIER DRIVE WARNING
   "Carrier_33_Status" AT %IW2000 : Word;   // CARRIER STATUS WORD
   "Carrier_33_Status.0" AT %I2000.0 : Bool;   // HEARTBEAT
   "Carrier_33_Status.1" AT %I2000.1 : Bool;   // MANUAL
   "Carrier_33_Status.2" AT %I2000.2 : Bool;   // IN_AUTO
   "Carrier_33_Status.3" AT %I2000.3 : Bool;   // POSITIONING_COMPLETE
   "Carrier_33_Status.4" AT %I2000.4 : Bool;   // PRODUCTION HOLD
   "Carrier_33_Status.5" AT %I2000.5 : Bool;   // CARRIER MOVING FORWARD
   "Carrier_33_Status.6" AT %I2000.6 : Bool;   // CARRIER MOVING REVERSE
   "Carrier_33_Status.7" AT %I2000.7 : Bool;   // CARRIER FAULT
   "Carrier_33_Status.8" AT %I2001.0 : Bool;   // CRASH DETECT TRIPPED
   "Carrier_33_Status.9" AT %I2001.1 : Bool;